// TIA Portal project "Inteligenta_szklarnia" (V15.1) (continued)

screen "tryb_automatyczny" 800x480
   IOField "I/O field_1" at 100,354 size 57x40; FormatPattern 99.9
      ProcessValue <- "Wejscia_HMI_Temperatura"
   Button "Button_1" at 750,0 size 50x50; TextOff 'WRÓĆ'; PictureOff "Back_arrow"
      on Click: function_efd93a16()
   Button "Button_2" at 417,418 size 371x53; TextOff 'ZATWIERDŹ'
      on Click: ActivateScreen("praca", 0)
   Bar "Bar_1" at 14,103 size 70x275; MinimumValue 0; MaximumValue 45
      ProcessValue <- "temperatura_ustawiona_man"
   TextField "Text field_2" at 15,60 size 132x23; Text 'TEMPERATURA'
   Bar "Bar_2" at 217,108 size 70x275; MinimumValue 0; MaximumValue 100
      ProcessValue <- "wilgotnosc_powietrza_man"
   TextField "Text field_3" at 205,61 size 122x42; Text 'WOLGOTNOŚĆ POWIETRZA WILGOTNOŚĆ POWIETRZA'
   Button "Button_3" at 90,119 size 75x45; TextOff '+ / +0.5 °C'
      on Press: function_dd21b452("temperatura_ustawiona_man", 0.5)
   Button "Button_7" at 89,177 size 75x45; TextOff '- / -0.5 °C'
      on Press: function_b9b71300("temperatura_ustawiona_man", 0.5)
   IOField "I/O field_2" at 100,276 size 62x40; FormatPattern 99.9
      ProcessValue <- "temperatura_ustawiona_man"
   TextField "Text field_11" at 155,285 size 23x22; Text '°C'
   TextField "Text field_9" at 155,358 size 23x22; Text '°C'
   Bar "Bar_4" at 417,105 size 70x275; MinimumValue 0; MaximumValue 100
      ProcessValue <- "wilgotnosc_gleby_man"
   TextField "Text field_10" at 404,58 size 122x42; Text 'WOLGOTNOŚĆ GLEBY WILGOTNOŚĆ GLEBY'
   Button "Button_8" at 496,125 size 65x40; TextOff '+ / +2%'
      on Click: function_dd21b452("wilgotnosc_gleby_man", 2)
   Button "Button_9" at 497,177 size 65x40; TextOff '- / -2%'
      on Click: function_b9b71300("wilgotnosc_gleby_man", 2)
   IOField "I/O field_5" at 508,276 size 62x40; FormatPattern 999
      ProcessValue <- "wilgotnosc_gleby_man"
   IOField "I/O field_6" at 508,346 size 62x40; FormatPattern 999
      ProcessValue <- "Parametry_Wilgotność_gleby"
   TextField "Text field_12" at 493,264 size 101x22; Text 'USTAWIONA'
   TextField "Text field_13" at 497,335 size 86x22; Text 'AKTUALNA'
   TextField "Text field_14" at 547,285 size 23x22; Text '%'
   TextField "Text field_15" at 547,356 size 23x22; Text '%'
   Button "Button_10" at 298,125 size 65x40; TextOff '+ / +5%'
      on Click: function_dd21b452("wilgotnosc_powietrza_man", 5)
   Button "Button_11" at 298,177 size 65x40; TextOff '- / -5%'
      on Click: function_b9b71300("wilgotnosc_powietrza_man", 5)
   IOField "I/O field_4" at 305,277 size 66x40; FormatPattern 999
      ProcessValue <- "wilgotnosc_powietrza_man"
   IOField "I/O field_7" at 307,349 size 62x40; FormatPattern 999
      ProcessValue <- "Parametry_Wilgotność_powietrza"
   TextField "Text field_16" at 292,264 size 101x22; Text 'USTAWIONA'
   TextField "Text field_17" at 294,335 size 86x22; Text 'AKTUALNA'
   TextField "Text field_18" at 346,286 size 23x22; Text '%'
   TextField "Text field_19" at 346,357 size 23x22; Text '%'
   Button "Button_14" at 3,1 size 43x43; TextOff 'DOM'; PictureOff "home_1"
      on Click: ActivateScreen("Root screen", 0)
   TextField "Text field_4" at 38,424 size 128x23; Text 'SYSTEM OKIEN'
   Switch "Switch_1" at 198,418 size 185x35; TextOn 'ON'; CaptionText 'Switch'; TextOff 'OFF'
      ProcessValue <- "system_okien"
   GraphicView "Graphic view_1" at 150,60 size 40x40; Picture "Thermometer_icon"
   GraphicView "Graphic view_2" at 330,61 size 40x40; Picture "sensor_4212519"
   TextField "Text field_5" at 93,334 size 86x22; Text 'AKTUALNA'
   TextField "Text field_6" at 90,262 size 101x22; Text 'USTAWIONA'
   GraphicView "Graphic view_3" at 526,61 size 40x40; Picture "soil-sensor_11298794"
   TextField "Text field_1" at 250,4 size 288x34; Text 'TRYB AUTOMATYCZNY'
   Bar "Bar_3" at 620,105 size 70x275; MinimumValue 0; MaximumValue 1500
      ProcessValue <- "wilgotnosc_gleby_man"
   TextField "Text field_7" at 604,53 size 161x42; Text 'WOLGOTNOŚĆ GLEBY NASŁONECZNIENIE'
   GraphicView "Graphic view_4" at 725,79 size 40x40; Picture "sensor_4212513"
   Button "Button_4" at 696,125 size 65x40; TextOff '+ +25 W m'
      on Click: function_dd21b452("naslonecznienie_man", 25)
   Button "Button_5" at 697,177 size 65x40; TextOff '- -25 W m'
      on Click: function_b9b71300("naslonecznienie_man", 25)
   IOField "I/O field_3" at 708,276 size 62x40; FormatPattern 999
      ProcessValue <- "naslonecznienie_man"
   TextField "Text field_8" at 693,264 size 101x22; Text 'USTAWIONA'
   IOField "I/O field_8" at 711,347 size 62x40; FormatPattern 999
      ProcessValue <- "Parametry_Czujnik_światła"
   TextField "Text field_20" at 697,335 size 86x22; Text 'AKTUALNA'
   TextField "Text field_21" at 747,285 size 23x22; Text '%'
   TextField "Text field_22" at 747,356 size 23x22; Text '%'
   TextField "Text field_23" at 751,143 size 32x18; Text '2'
   TextField "Text field_24" at 748,196 size 32x18; Text '2'
*)

(* ===== HMI "HMI_RT_3" =====
system functions are stored by id; their names below are inferred from use
connection "HMI_Connection_4": ETHERNET, SMART_S7_1200_OMS

HMI tags "Default tag table"
   "Tag_ScreenNumber" : UInt, internal

HMI tags "wyjsciaPLC"
   "Alarm_ostrzegwaczy" : Bool = PLC Alarm_ostrzegwaczy AT %Q0.5, 100 ms
   "Grzałka" : Bool = PLC Grzałka AT %Q0.0, 100 ms
   "Pompa_wodna" : Bool = PLC Pompa_wodna AT %Q0.2, 100 ms
   "Rolety_otwieranie" : Bool = PLC Rolety_otwieranie AT %Q0.3, 100 ms
   "Rolety_zamykanie" : Bool = PLC Rolety_zamykanie AT %Q0.4, 100 ms
   "Siłownik_okien_otwieranie" : Bool = PLC Siłownik_okien_otwieranie AT %Q0.6, 100 ms
   "Siłownik_okien_zamykanie" : Bool = PLC Siłownik_okien_zamykanie AT %Q0.7, 100 ms
   "Wentylator" : Bool = PLC Wentylator AT %Q0.1, 100 ms
   "Tag_ScreenNumber(1)" : DInt = PLC Tag_ScreenNumber AT %MD0, 500 ms
   "Parametry_Czujnik_światła" : Int = PLC Parametry.Czujnik_światła, 500 ms
   "Parametry_temeratura" : Real = PLC Parametry.temeratura, 500 ms
   "Parametry_Czujnik_wiatru" : Int = PLC Parametry.Czujnik_wiatru, 500 ms
   "Parametry_Wilgotność_powietrza" : Int = PLC Parametry.Wilgotność_powietrza, 500 ms
   "Parametry_czujnik_CO2" : Int = PLC Parametry.czujnik_CO2, 500 ms
   "Parametry_Wilgotność_gleby" : Int = PLC Parametry.Wilgotność_gleby, 500 ms
   "Wejscia_HMI_Temperatura" : Real = PLC Wejscia_HMI.Temperatura, 500 ms
   "Parametry_stopien_zasloniecia_rolet" : Int = PLC Parametry.stopien_zasloniecia_rolet, 1 s
   "Wejscia_HMI_Zaciemnienie" : Int = PLC Wejscia_HMI.Zaciemnienie, 1 s
   "Receptury_nazwa{0}" : String[254] = PLC Receptury.nazwa[0], 1 s
   "Receptury_nazwa{1}" : String[254] = PLC Receptury.nazwa[1], 1 s
   "Receptury_nazwa{2}" : String[254] = PLC Receptury.nazwa[2], 1 s
   "Receptury_nazwa{3}" : String[254] = PLC Receptury.nazwa[3], 1 s
   "Receptury_nazwa{4}" : String[254] = PLC Receptury.nazwa[4], 1 s
   "Receptury_nazwa{5}" : String[254] = PLC Receptury.nazwa[5], 1 s
   "naslonecznienie_man" : Int = PLC Wejscia_HMI.naslonecznienie_manual, 1 s

HMI tags "USTAWIENIA_HMI"
   "temperatura_ustawiona_man" : Real, internal
   "stopien_otwarcia_okien_man" : Real, internal
   "wilgotnosc_powietrza_man" : Real, internal
   "wilgotnosc_gleby_man" : Real, internal
   "nazwa_receptury" : WString[10], internal
   "system_okien" : Bool, internal
   "AlwaysTRUE" : Bool = PLC AlwaysTRUE AT %M1.2, 1 s

screen "Root screen" 800x480, template "Template_1"
   on GenerateScreen: SetTag("Tag_ScreenNumber", 1)
   Button "Button_3" at 10,270 size 300x90; TextOff 'ZAPISZ NOWĄ RECEPTURĘ'
      on Click: ActivateScreen("zapisz_recepture", 0)
   Button "Button_1" at 10,170 size 300x90; TextOff 'TRYB MANUALNY'
      on Click: ActivateScreen("tryb_manualny", 0)
   Button "Button_2" at 10,70 size 301x90; TextOff 'TRYB AUTOMATYCZNY'
      on Click: ActivateScreen("tryb_automatyczny", 0)
   TextField "Text field_2" at 32,2 size 738x63; Text 'AUTOMATYCZNA SZKLARNIA'
   GraphicView "Graphic view_1" at 370,70 size 392x338; Picture "garden-tools-graphic-clipart-design-free-png"
   Button "Button_4" at 10,370 size 301x90; TextOff 'WYBIERZ RECEPTURĘ'
      on Click: ActivateScreen("wybierz_recepture", 0)
   TextField "Text field_1" at 117,454 size 235x26; Text 'Tego przycisku w symulacji nie widac ale nie chciałem uswac jakby jednak był potrzebny xd'
      Visibility <- "AlwaysTRUE"

screen "zapisz_recepture" 800x480
   TextField "Text field_1" at 282,4 size 253x34; Text 'ZAPISZ RECEPTURE / ZAPISZ RECEPTURĘ'
   Button "Button_1" at 750,0 size 50x50; TextOff 'WRÓĆ'; PictureOff "Back_arrow"
      on Click: function_efd93a16()
   Button "Button_2" at 406,414 size 371x53; TextOff 'ZATWIERDŹ'
      on Click: ActivateScreen("praca", 0)
   Bar "Bar_1" at 17,122 size 70x314; MinimumValue 0; MaximumValue 45
      ProcessValue <- "temperatura_ustawiona_man"
   TextField "Text field_2" at 30,64 size 132x23; Text 'TEMPERATURA'
   Bar "Bar_2" at 223,133 size 54x113; MinimumValue 0; MaximumValue 100
      ProcessValue <- "wilgotnosc_powietrza_man"
   TextField "Text field_3" at 231,45 size 122x42; Text 'WOLGOTNOŚĆ POWIETRZA'
   Button "Button_3" at 115,140 size 73x45; TextOff '+ / +0.5 °C'
      on Press: function_dd21b452("temperatura_ustawiona_man", 0.5)
   Button "Button_7" at 115,201 size 73x45; TextOff '- / -0.5 °C'
      on Press: function_b9b71300("temperatura_ustawiona_man", 0.5)
   TextField "Text field_8" at 93,325 size 109x42; Text 'ustawiona wartość USTAWIONA'
   IOField "I/O field_2" at 106,365 size 62x40; FormatPattern 99.9
      ProcessValue <- "temperatura_ustawiona_man"
   TextField "Text field_11" at 156,367 size 37x37; Text '°C'
   Bar "Bar_4" at 225,346 size 57x127; MinimumValue 0; MaximumValue 100
      ProcessValue <- "wilgotnosc_gleby_man"
   TextField "Text field_10" at 229,254 size 122x42; Text 'WOLGOTNOŚĆ GLEBY'
   Button "Button_8" at 230,300 size 40x40; TextOff '+'
      on Click: function_dd21b452("wilgotnosc_gleby_man", 2)
   Button "Button_9" at 318,300 size 40x40; TextOff '-'
      on Click: function_b9b71300("wilgotnosc_gleby_man", 2)
   IOField "I/O field_5" at 291,401 size 62x40; FormatPattern 999
      ProcessValue <- "wilgotnosc_gleby_man"
   TextField "Text field_12" at 285,384 size 83x20; Text 'USTAWIONA'
   TextField "Text field_14" at 338,404 size 30x29; Text '%'
   Button "Button_10" at 223,87 size 40x40; TextOff '+'
      on Click: function_dd21b452("wilgotnosc_powietrza_man", 5)
   Button "Button_11" at 311,87 size 40x40; TextOff '-'
      on Click: function_b9b71300("wilgotnosc_powietrza_man", 5)
   IOField "I/O field_4" at 291,180 size 62x40; FormatPattern 999
      ProcessValue <- "wilgotnosc_powietrza_man"
   TextField "Text field_16" at 288,167 size 83x20; Text 'USTAWIONA'
   TextField "Text field_18" at 342,184 size 30x29; Text '%'
   Button "Button_14" at 3,1 size 43x43; TextOff 'DOM'; PictureOff "home_1"
      on Click: ActivateScreen("Root screen", 0)
   TextField "Text field_4" at 529,47 size 128x23; Text 'SYSTEM OKIEN'
   Switch "Switch_1" at 503,78 size 185x35; TextOn 'ON'; CaptionText 'Switch'; TextOff 'OFF'
      ProcessValue <- "system_okien"
   IOField "I/O field_1" at 426,311 size 328x81; FormatPattern ????????????????????
      ProcessValue <- "nazwa_receptury"
   TextField "Text field_7" at 406,273 size 380x37; Text 'WPISZ NAZWĘ RECEPTURY'
   GraphicView "Graphic view_1" at 385,338 size 36x30; Picture "Graphic_4"
   GraphicView "Graphic view_2" at 753,338 size 36x30; Picture "Graphic_5"
   TextField "Text field_9" at 387,146 size 161x61; Text 'STOPIEŃ OTWARCIA OKIEN ŚREDNIE NASŁONECZNIENIE'
   Bar "Bar_6" at 404,213 size 373x52; MinimumValue 0; MaximumValue 1500
      ProcessValue <- "naslonecznienie_man"
   Button "Button_4" at 697,145 size 80x50; TextOff '+ / -'
      on Click: function_b9b71300("naslonecznienie_man", 5)
   Button "Button_5" at 589,145 size 80x50; TextOff '- / +'
      on Press: function_dd21b452("naslonecznienie_man", 5)

screen "tryb_manualny" 800x480
   Button "Button_2" at 355,415 size 431x53; TextOff 'ZATWIERDŹ'
      on Click: ActivateScreen("praca", 0)
   TextField "Text field_1" at 282,4 size 223x34; Text 'TRYB MANUALNY'
   Bar "Bar_1" at 181,300 size 60x172; MinimumValue 0; MaximumValue 45
      ProcessValue <- "Parametry_temeratura"
   TextField "Text field_2" at 188,267 size 132x23; Text 'TEMPERATURA'
   Bar "Bar_2" at 181,93 size 60x160; MinimumValue 0; MaximumValue 100
      ProcessValue <- "Parametry_Wilgotność_powietrza"
   TextField "Text field_3" at 198,45 size 122x42; Text 'WOLGOTNOŚĆ POWIETRZA WILGOTNOŚĆ POWIETRZA'
   Bar "Bar_3" at 576,166 size 170x52; MinimumValue 0
      ProcessValue <- "stopien_otwarcia_okien_man"
   TextField "Text field_4" at 576,43 size 186x61; Text 'STOPIEŃ OTWARCIA OKIEN STOPIEŃ OTWARCIA OKIEN'
   IOField "I/O field_1" at 244,368 size 95x40; FormatPattern 99.9
      ProcessValue <- "Wejscia_HMI_Temperatura"
   Bar "Bar_4" at 8,93 size 60x160; MinimumValue 0; MaximumValue 100
      ProcessValue <- "Parametry_Wilgotność_gleby"
   Button "Button_4" at 406,253 size 80x60; TextOff 'PODLEWANIE'
      on Click: InvertBit("Pompa_wodna")
   Button "Button_5" at 536,253 size 80x60; TextOff 'GRZANIE'
      on Click: InvertBit("Grzałka")
   Button "Button_6" at 666,253 size 80x60; TextOff 'WENTYLACJA'
      on Click: InvertBit("Wentylator")
   GraphicView "Graphic view_1" at 675,320 size 60x60; Picture "fan_4829316"
      Visibility <- "Wentylator"
   GraphicView "Graphic view_6" at 545,320 size 60x60; Picture "heater_4463010"
      Visibility <- "Grzałka"
   GraphicView "Graphic view_7" at 415,320 size 60x60; Picture "irrigation_18631825"
      Visibility <- "Pompa_wodna"
   GraphicView "Graphic view_9" at 676,320 size 60x60; Picture "fan_off"
      Visibility <- "Wentylator"
   GraphicView "Graphic view_10" at 546,320 size 60x60; Picture "heater_off"
      Visibility <- "Grzałka"
   GraphicView "Graphic view_11" at 415,320 size 60x60; Picture "irrigation_off"
      Visibility <- "Pompa_wodna"
   TextField "Text field_10" at 18,45 size 122x42; Text 'WOLGOTNOŚĆ GLEBY WILGOTNOŚĆ GLEBY'
   IOField "I/O field_3" at 760,171 size 33x36; FormatPattern 9
      ProcessValue <- "stopien_otwarcia_okien_man"
   IOField "I/O field_6" at 70,148 size 62x40; FormatPattern 999
      ProcessValue <- "Parametry_Wilgotność_gleby"
   TextField "Text field_15" at 115,152 size 35x34; Text '%'
   IOField "I/O field_7" at 252,151 size 62x40; FormatPattern 999
      ProcessValue <- "Parametry_Wilgotność_powietrza"
   TextField "Text field_19" at 294,154 size 35x34; Text '%'
   Button "Button_12" at 576,99 size 50x50; TextOff '+'
      on Click: function_dd21b452("stopien_otwarcia_okien_man", 1)
   Button "Button_13" at 696,98 size 50x50; TextOff '-'
      on Click: function_b9b71300("stopien_otwarcia_okien_man", 1)
   Button "Button_14" at 3,1 size 43x43; TextOff 'DOM'; PictureOff "home_1"
      on Click: ActivateScreen("Root screen", 0)
   Button "Button_1" at 750,0 size 50x50; TextOff 'Text'; PictureOff "Back_arrow"
      on Click: function_efd93a16()
   TextField "Text field_9" at 293,369 size 35x34; Text '°C'
   Circle "Circle_1" at 386,336 size 25x25
      Visibility <- "Pompa_wodna"
   Circle "Circle_4" at 386,336 size 25x25
      Visibility <- "Pompa_wodna"
   Circle "Circle_2" at 511,336 size 25x25
      Visibility <- "Grzałka"
   Circle "Circle_5" at 511,336 size 25x25
      Visibility <- "Grzałka"
   Circle "Circle_3" at 639,336 size 25x25
      Visibility <- "Wentylator"
   Circle "Circle_6" at 639,336 size 25x25
      Visibility <- "Wentylator"
   Bar "Bar_5" at 10,300 size 60x172; MinimumValue 0; MaximumValue 1500
      ProcessValue <- "Parametry_Czujnik_światła"
   TextField "Text field_5" at 3,268 size 161x23; Text 'TEMPERATURA / NASŁONECZNIENIE'
   IOField "I/O field_2" at 70,368 size 95x40; FormatPattern 9999
      ProcessValue <- "Parametry_Czujnik_światła"
   TextField "Text field_6" at 127,356 size 35x64; Text '°C W m'
   TextField "Text field_7" at 152,391 size 31x17; Text '2'
   TextField "Text field_8" at 348,43 size 206x61; Text 'STOPIEŃ OTWARCIA OKIEN STOPIEŃ ZASŁONIENIA ROLET'
   Bar "Bar_6" at 366,166 size 170x52; MinimumValue 0; MaximumValue 100
      ProcessValue <- "naslonecznienie_man"
   Button "Button_3" at 456,98 size 80x50; TextOff '+ / ODSŁOŃ'
      on Click: function_b9b71300("naslonecznienie_man", 5)
   Button "Button_7" at 366,98 size 80x50; TextOff '- / ZASŁOŃ'
      on Press: function_dd21b452("naslonecznienie_man", 5)

screen "wybierz_recepture" 800x480
   TextField "Text field_2" at 257,4 size 280x34; Text 'WYBIERZ RECEPTURE / WYBIERZ RECEPTURĘ'
   Button "Button_1" at 750,0 size 50x50; TextOff 'WRÓĆ'; PictureOff "Back_arrow"
      on Click: function_efd93a16()
   Button "Button_14" at 3,1 size 43x43; TextOff 'DOM'; PictureOff "home_1"
      on Click: ActivateScreen("Root screen", 0)
   TextField "Text field_1" at 18,52 size 23x39; Text '1'
   TextField "Text field_3" at 18,108 size 23x39; Text '2'
   TextField "Text field_4" at 18,169 size 23x39; Text '3'
   TextField "Text field_5" at 18,231 size 23x39; Text '4'
   TextField "Text field_6" at 18,290 size 23x39; Text '5'
   TextField "Text field_7" at 18,351 size 23x39; Text '6'
   Button "Button_2" at 13,415 size 775x55; TextOff '-ZATWIERDŹ-'
      on Click: ActivateScreen("praca", 0)
   Button "Button_3" at 720,68 size 60x60; TextOff 'Text'; PictureOff "Double_up_arrow"
   Button "Button_4" at 720,162 size 60x60; TextOff 'Text'; PictureOff "Double_down_arrow"
   Button "Button_5" at 708,326 size 83x64; TextOff 'USUŃ'
   IOField "I/O field_1" at 90,58 size 243x32; FormatPattern ????????????????????
      ProcessValue <- "Receptury_nazwa{0}"
   IOField "I/O field_2" at 90,115 size 241x32; FormatPattern ????????????????????
      ProcessValue <- "Receptury_nazwa{1}"
   IOField "I/O field_3" at 90,176 size 267x32; FormatPattern ????????????????????
      ProcessValue <- "Receptury_nazwa{2}"
   IOField "I/O field_4" at 90,238 size 264x32; FormatPattern ????????????????????
      ProcessValue <- "Receptury_nazwa{3}"
   IOField "I/O field_5" at 90,294 size 230x32; FormatPattern ????????????????????
      ProcessValue <- "Receptury_nazwa{4}"
   IOField "I/O field_6" at 90,358 size 506x32; FormatPattern ????????????????????
      ProcessValue <- "Receptury_nazwa{5}"

screen "praca" 800x480
   GraphicView "Graphic view_2" at 28,217 size 100x100; Picture "Thermometer_icon"
   GraphicView "Graphic view_4" at 276,362 size 100x100; Picture "soil-sensor_11298794"
   GraphicView "Graphic view_3" at 28,74 size 100x100; Picture "sensor_4212513"
   GraphicView "Graphic view_5" at 276,75 size 100x100; Picture "sensor_4212519"
   GraphicView "Graphic view_1" at 559,362 size 100x100; Picture "fan_4829316"
      Visibility <- "Wentylator"
   GraphicView "Graphic view_6" at 560,217 size 100x100; Picture "heater_4463010"
      Visibility <- "Grzałka"
   GraphicView "Graphic view_7" at 560,75 size 100x100; Picture "irrigation_18631825"
      Visibility <- "Pompa_wodna"
   GraphicView "Graphic view_8" at 28,362 size 100x100; Picture "anemometer_1113716"
   GraphicView "Graphic view_9" at 560,362 size 100x100; Picture "fan_off"
      Visibility <- "Wentylator"
   GraphicView "Graphic view_10" at 561,217 size 100x100; Picture "heater_off"
      Visibility <- "Grzałka"
   GraphicView "Graphic view_11" at 561,75 size 100x100; Picture "irrigation_off"
      Visibility <- "Pompa_wodna"
   GraphicView "Graphic view_12" at 276,217 size 100x100; Picture "sensor_2828470"
   TextField "Text field_1" at 54,52 size 204x23; Text 'INSOLATION / NASŁONECZNIENIE / SONNENEINSTRAHLUNG'
   TextField "Text field_2" at 67,194 size 132x23; Text 'TEMPERATURA'
   TextField "Text field_3" at 46,334 size 166x23; Text 'SZYBKOŚĆ WIATRU'
   TextField "Text field_4" at 349,194 size 123x23; Text 'STĘŻENIE CO2'
   TextField "Text field_5" at 294,50 size 223x23; Text 'WILGOTNOŚĆ POWIETRZA'
   TextField "Text field_6" at 321,339 size 175x23; Text 'WILGOTNOŚĆ GLEBY'
   TextField "Text field_7" at 626,46 size 116x23; Text 'PODLEWANIE'
   TextField "Text field_8" at 643,192 size 80x23; Text 'GRZANIE'
   TextField "Text field_9" at 626,330 size 117x23; Text 'WENTYLACJA'
   TextField "Text field_10" at 282,4 size 256x34; Text 'PODGLĄD NA ŻYWO'
   Button "Button_1" at 750,0 size 50x50; TextOff 'WRÓĆ'; PictureOff "Back_arrow"
      on Click: function_efd93a16()
   Button "Button_2" at 3,1 size 43x43; TextOff 'DOM'; PictureOff "home_1"
      on Click: ActivateScreen("Root screen", 0)
   IOField "I/O field_2" at 120,233 size 97x65; FormatPattern 99.99
      ProcessValue <- "Parametry_temeratura"
   IOField "I/O field_3" at 136,383 size 70x65; FormatPattern 999
      ProcessValue <- "Parametry_Czujnik_wiatru"
   IOField "I/O field_5" at 377,235 size 83x65; FormatPattern 9999
      ProcessValue <- "Parametry_czujnik_CO2"
   TextField "Text field_11" at 214,241 size 46x46; Text '°C'
   IOField "I/O field_4" at 406,95 size 69x65; FormatPattern 999
      ProcessValue <- "Parametry_Wilgotność_powietrza"
   IOField "I/O field_6" at 406,384 size 68x65; FormatPattern 999
      ProcessValue <- "Parametry_Wilgotność_gleby"
   TextField "Text field_12" at 472,106 size 47x46; Text '%'
   TextField "Text field_13" at 472,396 size 47x46; Text '%'
   TextField "Text field_14" at 219,90 size 47x72; Text 'W m²'
   IOField "I/O field_1" at 119,109 size 101x32; FormatPattern 99999
      ProcessValue <- "Parametry_Czujnik_światła"
   TextField "Text field_15" at 210,376 size 52x72; Text 'Km h'
   Circle "Circle_1" at 695,101 size 48x48
      Visibility <- "Pompa_wodna"
   Circle "Circle_2" at 695,243 size 48x48
      Visibility <- "Grzałka"
   TextField "Text field_16" at 472,242 size 69x39; Text 'ppm'
   Circle "Circle_4" at 695,101 size 48x48
      Visibility <- "Pompa_wodna"
   Circle "Circle_5" at 695,243 size 48x48
      Visibility <- "Grzałka"
   Circle "Circle_3" at 695,385 size 48x48
      Visibility <- "Wentylator"
   Circle "Circle_6" at 695,385 size 48x48
      Visibility <- "Wentylator"

screen "tryb_automatyczny" 800x480
   IOField "I/O field_1" at 100,354 size 57x40; FormatPattern 99.9
      ProcessValue <- "Wejscia_HMI_Temperatura"
   Button "Button_1" at 750,0 size 50x50; TextOff 'WRÓĆ'; PictureOff "Back_arrow"
      on Click: function_efd93a16()
   Button "Button_2" at 417,418 size 371x53; TextOff 'ZATWIERDŹ'
      on Click: ActivateScreen("praca", 0)
   Bar "Bar_1" at 14,103 size 70x275; MinimumValue 0; MaximumValue 45
      ProcessValue <- "temperatura_ustawiona_man"
   TextField "Text field_2" at 15,60 size 132x23; Text 'TEMPERATURA'
   Bar "Bar_2" at 217,108 size 70x275; MinimumValue 0; MaximumValue 100
      ProcessValue <- "wilgotnosc_powietrza_man"
   TextField "Text field_3" at 205,61 size 122x42; Text 'WOLGOTNOŚĆ POWIETRZA WILGOTNOŚĆ POWIETRZA'
   Button "Button_3" at 90,119 size 75x45; TextOff '+ / +0.5 °C'
      on Press: function_dd21b452("temperatura_ustawiona_man", 0.5)
   Button "Button_7" at 89,177 size 75x45; TextOff '- / -0.5 °C'
      on Press: function_b9b71300("temperatura_ustawiona_man", 0.5)
   IOField "I/O field_2" at 100,276 size 62x40; FormatPattern 99.9
      ProcessValue <- "temperatura_ustawiona_man"
   TextField "Text field_11" at 155,285 size 23x22; Text '°C'
   TextField "Text field_9" at 155,358 size 23x22; Text '°C'
   Bar "Bar_4" at 417,105 size 70x275; MinimumValue 0; MaximumValue 100
      ProcessValue <- "wilgotnosc_gleby_man"
   TextField "Text field_10" at 404,58 size 122x42; Text 'WOLGOTNOŚĆ GLEBY WILGOTNOŚĆ GLEBY'
   Button "Button_8" at 496,125 size 65x40; TextOff '+ / +2%'
      on Click: function_dd21b452("wilgotnosc_gleby_man", 2)
   Button "Button_9" at 497,177 size 65x40; TextOff '- / -2%'
      on Click: function_b9b71300("wilgotnosc_gleby_man", 2)
   IOField "I/O field_5" at 508,276 size 62x40; FormatPattern 999
      ProcessValue <- "wilgotnosc_gleby_man"
   IOField "I/O field_6" at 508,346 size 62x40; FormatPattern 999
      ProcessValue <- "Parametry_Wilgotność_gleby"
   TextField "Text field_12" at 493,264 size 101x22; Text 'USTAWIONA'
   TextField "Text field_13" at 497,335 size 86x22; Text 'AKTUALNA'
   TextField "Text field_14" at 547,285 size 23x22; Text '%'
   TextField "Text field_15" at 547,356 size 23x22; Text '%'
   Button "Button_10" at 298,125 size 65x40; TextOff '+ / +5%'
      on Click: function_dd21b452("wilgotnosc_powietrza_man", 5)
   Button "Button_11" at 298,177 size 65x40; TextOff '- / -5%'
      on Click: function_b9b71300("wilgotnosc_powietrza_man", 5)
   IOField "I/O field_4" at 305,277 size 66x40; FormatPattern 999
      ProcessValue <- "wilgotnosc_powietrza_man"
   IOField "I/O field_7" at 307,349 size 62x40; FormatPattern 999
      ProcessValue <- "Parametry_Wilgotność_powietrza"
   TextField "Text field_16" at 292,264 size 101x22; Text 'USTAWIONA'
   TextField "Text field_17" at 294,335 size 86x22; Text 'AKTUALNA'
   TextField "Text field_18" at 346,286 size 23x22; Text '%'
   TextField "Text field_19" at 346,357 size 23x22; Text '%'
   Button "Button_14" at 3,1 size 43x43; TextOff 'DOM'; PictureOff "home_1"
      on Click: ActivateScreen("Root screen", 0)
   TextField "Text field_4" at 38,424 size 128x23; Text 'SYSTEM OKIEN'
   Switch "Switch_1" at 198,418 size 185x35; TextOn 'ON'; CaptionText 'Switch'; TextOff 'OFF'
      ProcessValue <- "system_okien"
   GraphicView "Graphic view_1" at 150,60 size 40x40; Picture "Thermometer_icon"
   GraphicView "Graphic view_2" at 330,61 size 40x40; Picture "sensor_4212519"
   TextField "Text field_5" at 93,334 size 86x22; Text 'AKTUALNA'
   TextField "Text field_6" at 90,262 size 101x22; Text 'USTAWIONA'
   GraphicView "Graphic view_3" at 526,61 size 40x40; Picture "soil-sensor_11298794"
   TextField "Text field_1" at 250,4 size 288x34; Text 'TRYB AUTOMATYCZNY'
   Bar "Bar_3" at 620,105 size 70x275; MinimumValue 0; MaximumValue 1500
      ProcessValue <- "wilgotnosc_gleby_man"
   TextField "Text field_7" at 604,53 size 161x42; Text 'WOLGOTNOŚĆ GLEBY NASŁONECZNIENIE'
   GraphicView "Graphic view_4" at 725,79 size 40x40; Picture "sensor_4212513"
   Button "Button_4" at 696,125 size 65x40; TextOff '+ +25 W m'
      on Click: function_dd21b452("naslonecznienie_man", 25)
   Button "Button_5" at 697,177 size 65x40; TextOff '- -25 W m'
      on Click: function_b9b71300("naslonecznienie_man", 25)
   IOField "I/O field_3" at 708,276 size 62x40; FormatPattern 999
      ProcessValue <- "naslonecznienie_man"
   TextField "Text field_8" at 693,264 size 101x22; Text 'USTAWIONA'
   IOField "I/O field_8" at 711,347 size 62x40; FormatPattern 999
      ProcessValue <- "Parametry_Czujnik_światła"
   TextField "Text field_20" at 697,335 size 86x22; Text 'AKTUALNA'
   TextField "Text field_21" at 747,285 size 23x22; Text '%'
   TextField "Text field_22" at 747,356 size 23x22; Text '%'
   TextField "Text field_23" at 751,143 size 32x18; Text '2'
   TextField "Text field_24" at 748,196 size 32x18; Text '2'

Template "Template_1" 800x480
   Button "Exit" at 671,429 size 71x50; TextOn 'Exit'; TextOff 'Exit'; PictureOn "ExitRuntime_KTP700_Basic_PN_TR"; PictureOff "ExitRuntime_KTP700_Basic_PN_TR"
      on Release: StopRuntime(0)
   Button "Alarms" at 524,429 size 71x50; TextOn 'Alarms'; TextOff 'Alarms'; PictureOn "AlarmDisplay_KTP700_Basic_PN_TR"; PictureOff "AlarmDisplay_KTP700_Basic_PN_TR"
      on Release: function_ef3f5d25("Alarm window_Unacknowledged", -1)
   Button "Start screen" at 169,429 size 71x50; TextOn 'Start screen'; TextOff 'Start screen'; PictureOn "NavigateHome_KTP700_Basic_PN_TR"; PictureOff "NavigateHome_KTP700_Basic_PN_TR"
      on Release: ActivateScreen("Root screen", 0)
      Visibility <- "AlwaysTRUE"
   Button "Language" at 377,429 size 71x50; TextOn 'Language'; TextOff 'Language'; PictureOn "ToggleLanguage_KTP700_Basic_PN_TR"; PictureOff "ToggleLanguage_KTP700_Basic_PN_TR"
      on Release: function_fb9197e8(-1)
*)

(* ===== HMI "HMI_RT_2" =====
system functions are stored by id; their names below are inferred from use
connection "HMI_Connection_3": ETHERNET, SMART_S7_1200_OMS

HMI tags "Default tag table"
   "Tag_ScreenNumber" : Int = PLC HMI.Numer_ekranu_HMI AT %MD0, 500 ms
   "AlwaysTRUE" : Bool = PLC AlwaysTRUE AT %M1.2, 1 s

HMI tags "Receptury"
   "Receptury_nazwa{0}" : String[254] = PLC Receptury.nazwa[0], 1 s
   "Receptury_nazwa{1}" : String[254] = PLC Receptury.nazwa[1], 1 s
   "Receptury_nazwa{2}" : String[254] = PLC Receptury.nazwa[2], 1 s
   "Receptury_nazwa{3}" : String[254] = PLC Receptury.nazwa[3], 1 s
   "Receptury_nazwa{4}" : String[254] = PLC Receptury.nazwa[4], 1 s
   "Receptury_nazwa{5}" : String[254] = PLC Receptury.nazwa[5], 1 s

HMI tags "USTAWIENIA_HMI"
   "nazwa_receptury" : WString[10], internal

HMI tags "Do_PLC"
   "System_okien_auto" : Bool = PLC HMI.System_okien_auto, 500 ms
   "Stopien_zasloniecia_rolet_manual" : Int = PLC HMI.Stopien_zasloniecia_rolet_manual, 100 ms
   "Przycisk_pompy_manual" : Bool = PLC HMI.Przycisk_pompa_manual AT %Q0.2, 100 ms
   "Przycisk_wentylacja_manual" : Bool = PLC HMI.Przycisk_wentylacja_manual AT %Q0.1, 100 ms
   "Przycisk_grzanie_manual" : Bool = PLC HMI.Przycisk_grzanie_manual AT %Q0.0, 100 ms
   "Stopien_otwarcia_okien_man" : Int = PLC HMI.Stopien_otwarcia_okien_manual AT %DB1.DBW0, 100 ms
   "Temperatura_auto" : Real = PLC HMI.Temperatura_auto, 500 ms
   "Naslonecznienie_auto" : Int = PLC HMI.Naslonecznienie_auto AT %DB1.DBW0, 500 ms
   "Wilgotnosc_powietrza_auto" : Int = PLC HMI.Wilgotnosc_powietrza_auto AT %DB1.DBW0, 500 ms
   "Wilgotnosc_gleby_auto" : Int = PLC HMI.Wilgotnosc_gleby_auto AT %DB1.DBW0, 500 ms
   "Przycisk_zatwierdz" : Bool = PLC HMI.Przycisk_zatwierdz AT %DB1.DBW0, 100 ms

HMI tags "Z_PLC"
   "Czujnik_wilgotności_powietrza" : Int = PLC Wejscia_PLC.Czujnik_wilgotności_powietrza, 500 ms
   "Czujnik_temeratury_wewnetrznej" : Real = PLC Wejscia_PLC.Temeratura_wewnetrzna, 500 ms
   "Czujnik_natezenia_światła" : Int = PLC Wejscia_PLC.Czujnik_natezenia_swiatła, 500 ms
   "Czujnik_wilgotności_gleby" : Int = PLC Wejscia_PLC.Czujnik_wilgotności_gleby, 500 ms
   "Czujnik_CO2" : Int = PLC Wejscia_PLC.Czujnik_CO2, 500 ms
   "Czujnik_wiatru" : Int = PLC Wejscia_PLC.Czujnik_wiatru, 500 ms
   "Stopien_zasloniecia_rolet" : Int = PLC Wejscia_PLC.Stopien_zasloniecia_rolet, 1 s

screen "Root screen" 800x480, template "Template_1"
   on GenerateScreen: SetTag("Tag_ScreenNumber", 0)
   Button "Button_3" at 10,270 size 300x90; TextOff 'ZAPISZ NOWĄ RECEPTURĘ'
      on Click: ActivateScreen("zapisz_recepture", 0)
   Button "Button_1" at 10,170 size 300x90; TextOff 'TRYB MANUALNY'
      on Click: ActivateScreen("tryb_manualny", 0)
   Button "Button_2" at 10,70 size 301x90; TextOff 'TRYB AUTOMATYCZNY'
      on Click: ActivateScreen("tryb_automatyczny", 0)
   TextField "Text field_2" at 32,2 size 738x63; Text 'AUTOMATYCZNA SZKLARNIA'
   GraphicView "Graphic view_1" at 370,70 size 392x338; Picture "garden-tools-graphic-clipart-design-free-png"
   Button "Button_4" at 10,370 size 301x90; TextOff 'WYBIERZ RECEPTURĘ'
      on Click: ActivateScreen("wybierz_recepture", 0)

screen "zapisz_recepture" 800x480
   on GenerateScreen: SetTag("Tag_ScreenNumber", 4)
   TextField "Text field_1" at 282,4 size 253x34; Text 'ZAPISZ RECEPTURE / ZAPISZ RECEPTURĘ'
   Button "Button_1" at 750,0 size 50x50; TextOff 'WRÓĆ'; PictureOff "Back_arrow"
      on Click: function_efd93a16()
   Button "Button_2" at 406,414 size 371x53; TextOff 'ZATWIERDŹ'
      on Click: ActivateScreen("praca", 0)
      on Press: function_b14e0dd5("Przycisk_zatwierdz", 0)
   Bar "Bar_1" at 17,122 size 70x314; MinimumValue 0; MaximumValue 45
      ProcessValue <- "Temperatura_auto"
   TextField "Text field_2" at 30,64 size 132x23; Text 'TEMPERATURA'
   Bar "Bar_2" at 223,133 size 54x113; MinimumValue 0; MaximumValue 100
      ProcessValue <- "Wilgotnosc_powietrza_auto"
   TextField "Text field_3" at 231,45 size 122x42; Text 'WOLGOTNOŚĆ POWIETRZA'
   Button "Button_3" at 115,140 size 73x45; TextOff '+ / +0.5 °C'
      on Press: function_dd21b452("Temperatura_auto", 0.5)
   Button "Button_7" at 115,201 size 73x45; TextOff '- / -0.5 °C'
      on Press: function_b9b71300("Temperatura_auto", 0.5)
   TextField "Text field_8" at 93,325 size 109x42; Text 'ustawiona wartość USTAWIONA'
   IOField "I/O field_2" at 106,365 size 62x40; FormatPattern 99.9
      ProcessValue <- "Temperatura_auto"
   TextField "Text field_11" at 156,367 size 37x37; Text '°C'
   Bar "Bar_4" at 225,346 size 57x127; MinimumValue 0; MaximumValue 100
      ProcessValue <- "Wilgotnosc_gleby_auto"
   TextField "Text field_10" at 229,254 size 122x42; Text 'WOLGOTNOŚĆ GLEBY'
   Button "Button_8" at 230,300 size 40x40; TextOff '+'
      on Click: function_dd21b452("Wilgotnosc_gleby_auto", 2)
   Button "Button_9" at 318,300 size 40x40; TextOff '-'
      on Click: function_b9b71300("Wilgotnosc_gleby_auto", 2)
   IOField "I/O field_5" at 291,401 size 62x40; FormatPattern 999
      ProcessValue <- "Wilgotnosc_gleby_auto"
   TextField "Text field_12" at 285,384 size 83x20; Text 'USTAWIONA'
   TextField "Text field_14" at 338,404 size 30x29; Text '%'
   Button "Button_10" at 223,87 size 40x40; TextOff '+'
      on Click: function_dd21b452("Wilgotnosc_powietrza_auto", 5)
   Button "Button_11" at 311,87 size 40x40; TextOff '-'
      on Click: function_b9b71300("Wilgotnosc_powietrza_auto", 5)
   IOField "I/O field_4" at 291,180 size 62x40; FormatPattern 999
      ProcessValue <- "Wilgotnosc_powietrza_auto"
   TextField "Text field_16" at 288,167 size 83x20; Text 'USTAWIONA'
   TextField "Text field_18" at 342,184 size 30x29; Text '%'
   Button "Button_14" at 3,1 size 43x43; TextOff 'DOM'; PictureOff "home_1"
      on Click: ActivateScreen("Root screen", 0)
   TextField "Text field_4" at 529,47 size 128x23; Text 'SYSTEM OKIEN'
   Switch "Switch_1" at 503,78 size 185x35; TextOn 'ON'; CaptionText 'Switch'; TextOff 'OFF'
      ProcessValue <- "System_okien_auto"
   IOField "I/O field_1" at 426,311 size 328x81; FormatPattern ????????????????????
      ProcessValue <- "nazwa_receptury"
   TextField "Text field_7" at 406,273 size 380x37; Text 'WPISZ NAZWĘ RECEPTURY'
   GraphicView "Graphic view_1" at 385,338 size 36x30; Picture "Graphic_4"
   GraphicView "Graphic view_2" at 753,338 size 36x30; Picture "Graphic_5"
   TextField "Text field_9" at 387,146 size 161x61; Text 'STOPIEŃ OTWARCIA OKIEN ŚREDNIE NASŁONECZNIENIE'
   Bar "Bar_6" at 404,213 size 373x52; MinimumValue 0; MaximumValue 1500
      ProcessValue <- "Stopien_zasloniecia_rolet_manual"
   Button "Button_4" at 697,145 size 80x50; TextOff '+ / -'
      on Click: function_b9b71300("Stopien_zasloniecia_rolet_manual", 5)
   Button "Button_5" at 589,145 size 80x50; TextOff '- / +'
      on Press: function_dd21b452("Stopien_zasloniecia_rolet_manual", 5)

screen "tryb_manualny" 800x480
   on GenerateScreen: SetTag("Tag_ScreenNumber", 2)
   TextField "Text field_1" at 282,4 size 223x34; Text 'TRYB MANUALNY'
   Bar "Bar_1" at 181,300 size 60x172; MinimumValue 0; MaximumValue 45
      ProcessValue <- "Czujnik_temeratury_wewnetrznej"
   TextField "Text field_2" at 188,267 size 132x23; Text 'TEMPERATURA'
   Bar "Bar_2" at 181,93 size 60x160; MinimumValue 0; MaximumValue 100
      ProcessValue <- "Czujnik_wilgotności_powietrza"
   TextField "Text field_3" at 198,45 size 122x42; Text 'WOLGOTNOŚĆ POWIETRZA WILGOTNOŚĆ POWIETRZA'
   Bar "Bar_3" at 576,166 size 170x52; MinimumValue 0
      ProcessValue <- "Stopien_otwarcia_okien_man"
   TextField "Text field_4" at 576,43 size 186x61; Text 'STOPIEŃ OTWARCIA OKIEN STOPIEŃ OTWARCIA OKIEN'
   IOField "I/O field_1" at 244,368 size 95x40; FormatPattern 99.9
      ProcessValue <- "Czujnik_temeratury_wewnetrznej"
   Bar "Bar_4" at 8,93 size 60x160; MinimumValue 0; MaximumValue 100
      ProcessValue <- "Czujnik_wilgotności_gleby"
   Button "Button_4" at 380,253 size 97x80; TextOff 'PODLEWANIE'
      on Click: InvertBit("Przycisk_pompy_manual")
   Button "Button_5" at 522,253 size 100x80; TextOff 'GRZANIE'
      on Click: InvertBit("Przycisk_grzanie_manual")
   Button "Button_6" at 671,253 size 100x80; TextOff 'WENTYLACJA'
      on Click: InvertBit("Przycisk_wentylacja_manual")
   GraphicView "Graphic view_1" at 681,356 size 76x80; Picture "fan_4829316"
      Visibility <- "Przycisk_wentylacja_manual"
   GraphicView "Graphic view_6" at 529,356 size 80x80; Picture "heater_4463010"
      Visibility <- "Przycisk_grzanie_manual"
   GraphicView "Graphic view_7" at 394,356 size 77x80; Picture "irrigation_18631825"
      Visibility <- "Przycisk_pompy_manual"
   GraphicView "Graphic view_9" at 682,356 size 76x80; Picture "fan_off"
      Visibility <- "Przycisk_wentylacja_manual"
   GraphicView "Graphic view_10" at 530,356 size 80x80; Picture "heater_off"
      Visibility <- "Przycisk_grzanie_manual"
   GraphicView "Graphic view_11" at 394,356 size 77x80; Picture "irrigation_off"
      Visibility <- "Przycisk_pompy_manual"
   TextField "Text field_10" at 18,45 size 122x42; Text 'WOLGOTNOŚĆ GLEBY WILGOTNOŚĆ GLEBY'
   IOField "I/O field_3" at 760,171 size 33x36; FormatPattern 9
      ProcessValue <- "Stopien_otwarcia_okien_man"
   IOField "I/O field_6" at 70,148 size 62x40; FormatPattern 999
      ProcessValue <- "Czujnik_wilgotności_gleby"
   TextField "Text field_15" at 115,152 size 35x34; Text '%'
   IOField "I/O field_7" at 252,151 size 62x40; FormatPattern 999
      ProcessValue <- "Czujnik_wilgotności_powietrza"
   TextField "Text field_19" at 294,154 size 35x34; Text '%'
   Button "Button_12" at 576,99 size 50x50; TextOff '+'
      on Click: function_dd21b452("Stopien_otwarcia_okien_man", 1)
   Button "Button_13" at 696,98 size 50x50; TextOff '-'
      on Click: function_b9b71300("Stopien_otwarcia_okien_man", 1)
   Button "Button_14" at 3,1 size 43x43; TextOff 'DOM'; PictureOff "home_1"
      on Click: ActivateScreen("Root screen", 0)
   Button "Button_1" at 750,0 size 50x50; TextOff 'Text'; PictureOff "Back_arrow"
      on Click: function_efd93a16()
   TextField "Text field_9" at 293,369 size 35x34; Text '°C'
   Circle "Circle_1" at 352,378 size 42x42
      Visibility <- "Przycisk_pompy_manual"
   Circle "Circle_4" at 352,378 size 42x42
      Visibility <- "Przycisk_pompy_manual"
   Circle "Circle_2" at 486,375 size 42x42
      Visibility <- "Przycisk_grzanie_manual"
   Circle "Circle_5" at 486,375 size 42x42
      Visibility <- "Przycisk_grzanie_manual"
   Circle "Circle_3" at 630,375 size 41x41
      Visibility <- "Przycisk_wentylacja_manual"
   Circle "Circle_6" at 630,375 size 41x41
      Visibility <- "Przycisk_wentylacja_manual"
   Bar "Bar_5" at 10,300 size 60x172; MinimumValue 0; MaximumValue 1500
      ProcessValue <- "Czujnik_natezenia_światła"
   TextField "Text field_5" at 3,268 size 161x23; Text 'TEMPERATURA / NASŁONECZNIENIE'
   IOField "I/O field_2" at 70,368 size 95x40; FormatPattern 9999
      ProcessValue <- "Czujnik_natezenia_światła"
   TextField "Text field_6" at 127,356 size 35x64; Text '°C W m'
   TextField "Text field_7" at 152,391 size 31x17; Text '2'
   TextField "Text field_8" at 348,43 size 205x61; Text 'STOPIEŃ OTWARCIA OKIEN STOPIEŃ ZASŁONIECIA ROLET'
   Bar "Bar_6" at 366,166 size 170x52; MinimumValue 0; MaximumValue 100
      ProcessValue <- "Stopien_zasloniecia_rolet_manual"
   Button "Button_3" at 456,98 size 80x50; TextOff '+ / ODSŁOŃ'
      on Click: function_b9b71300("Stopien_zasloniecia_rolet_manual", 5)
   Button "Button_7" at 366,98 size 80x50; TextOff '- / ZASŁOŃ'
      on Press: function_dd21b452("Stopien_zasloniecia_rolet_manual", 5)

screen "wybierz_recepture" 800x480
   on GenerateScreen: SetTag("Tag_ScreenNumber", 3)
   TextField "Text field_2" at 257,4 size 280x34; Text 'WYBIERZ RECEPTURE / WYBIERZ RECEPTURĘ'
   Button "Button_1" at 750,0 size 50x50; TextOff 'WRÓĆ'; PictureOff "Back_arrow"
      on Click: function_efd93a16()
   Button "Button_14" at 3,1 size 43x43; TextOff 'DOM'; PictureOff "home_1"
      on Click: ActivateScreen("Root screen", 0)
   TextField "Text field_1" at 18,52 size 23x39; Text '1'
   TextField "Text field_3" at 18,108 size 23x39; Text '2'
   TextField "Text field_4" at 18,169 size 23x39; Text '3'
   TextField "Text field_5" at 18,231 size 23x39; Text '4'
   TextField "Text field_6" at 18,290 size 23x39; Text '5'
   TextField "Text field_7" at 18,351 size 23x39; Text '6'
   Button "Button_2" at 13,415 size 775x55; TextOff '-ZATWIERDŹ-'
      on Click: ActivateScreen("praca", 0)
      on Press: function_b14e0dd5("Przycisk_zatwierdz", 0)
   Button "Button_3" at 720,68 size 60x60; TextOff 'Text'; PictureOff "Double_up_arrow"
   Button "Button_4" at 720,162 size 60x60; TextOff 'Text'; PictureOff "Double_down_arrow"
   Button "Button_5" at 708,326 size 83x64; TextOff 'USUŃ'
   IOField "I/O field_1" at 90,58 size 243x32; FormatPattern ????????????????????
      ProcessValue <- "Receptury_nazwa{0}"
   IOField "I/O field_2" at 90,115 size 241x32; FormatPattern ????????????????????
      ProcessValue <- "Receptury_nazwa{1}"
   IOField "I/O field_3" at 90,176 size 267x32; FormatPattern ????????????????????
      ProcessValue <- "Receptury_nazwa{2}"
   IOField "I/O field_4" at 90,238 size 264x32; FormatPattern ????????????????????
      ProcessValue <- "Receptury_nazwa{3}"
   IOField "I/O field_5" at 90,294 size 230x32; FormatPattern ????????????????????
      ProcessValue <- "Receptury_nazwa{4}"
   IOField "I/O field_6" at 90,358 size 506x32; FormatPattern ????????????????????
      ProcessValue <- "Receptury_nazwa{5}"

screen "praca" 800x480
   on GenerateScreen: SetTag("Tag_ScreenNumber", 5)
   GraphicView "Graphic view_2" at 28,217 size 100x100; Picture "Thermometer_icon"
   GraphicView "Graphic view_4" at 276,362 size 100x100; Picture "soil-sensor_11298794"
   GraphicView "Graphic view_3" at 28,74 size 100x100; Picture "sensor_4212513"
   GraphicView "Graphic view_5" at 276,75 size 100x100; Picture "sensor_4212519"
   GraphicView "Graphic view_1" at 559,362 size 100x100; Picture "fan_4829316"
      Visibility <- "Przycisk_wentylacja_manual"
   GraphicView "Graphic view_6" at 560,217 size 100x100; Picture "heater_4463010"
      Visibility <- "Przycisk_grzanie_manual"
   GraphicView "Graphic view_7" at 560,75 size 100x100; Picture "irrigation_18631825"
      Visibility <- "Przycisk_pompy_manual"
   GraphicView "Graphic view_8" at 28,362 size 100x100; Picture "anemometer_1113716"
   GraphicView "Graphic view_9" at 560,362 size 100x100; Picture "fan_off"
      Visibility <- "Przycisk_wentylacja_manual"
   GraphicView "Graphic view_10" at 561,217 size 100x100; Picture "heater_off"
      Visibility <- "Przycisk_grzanie_manual"
   GraphicView "Graphic view_11" at 561,75 size 100x100; Picture "irrigation_off"
      Visibility <- "Przycisk_pompy_manual"
   GraphicView "Graphic view_12" at 276,217 size 100x100; Picture "sensor_2828470"
   TextField "Text field_1" at 54,52 size 204x23; Text 'INSOLATION / NASŁONECZNIENIE / SONNENEINSTRAHLUNG'
   TextField "Text field_2" at 67,194 size 132x23; Text 'TEMPERATURA'
   TextField "Text field_3" at 46,334 size 166x23; Text 'SZYBKOŚĆ WIATRU'
   TextField "Text field_4" at 349,194 size 123x23; Text 'STĘŻENIE CO2'
   TextField "Text field_5" at 294,50 size 223x23; Text 'WILGOTNOŚĆ POWIETRZA'
   TextField "Text field_6" at 321,339 size 175x23; Text 'WILGOTNOŚĆ GLEBY'
   TextField "Text field_7" at 626,46 size 116x23; Text 'PODLEWANIE'
   TextField "Text field_8" at 643,192 size 80x23; Text 'GRZANIE'
   TextField "Text field_9" at 626,330 size 117x23; Text 'WENTYLACJA'
   TextField "Text field_10" at 282,4 size 256x34; Text 'PODGLĄD NA ŻYWO'
   Button "Button_1" at 750,0 size 50x50; TextOff 'WRÓĆ'; PictureOff "Back_arrow"
      on Click: function_efd93a16()
   Button "Button_2" at 3,1 size 43x43; TextOff 'DOM'; PictureOff "home_1"
      on Click: ActivateScreen("Root screen", 0)
   IOField "I/O field_2" at 120,233 size 97x65; FormatPattern 99.99
      ProcessValue <- "Czujnik_temeratury_wewnetrznej"
   IOField "I/O field_3" at 136,383 size 70x65; FormatPattern 999
      ProcessValue <- "Czujnik_wiatru"
   IOField "I/O field_5" at 377,235 size 83x65; FormatPattern 9999
      ProcessValue <- "Czujnik_CO2"
   TextField "Text field_11" at 214,241 size 46x46; Text '°C'
   IOField "I/O field_4" at 406,95 size 69x65; FormatPattern 999
      ProcessValue <- "Czujnik_wilgotności_powietrza"
   IOField "I/O field_6" at 406,384 size 68x65; FormatPattern 999
      ProcessValue <- "Czujnik_wilgotności_gleby"
   TextField "Text field_12" at 472,106 size 47x46; Text '%'
   TextField "Text field_13" at 472,396 size 47x46; Text '%'
   TextField "Text field_14" at 219,90 size 47x72; Text 'W m²'
   IOField "I/O field_1" at 119,109 size 101x32; FormatPattern 99999
      ProcessValue <- "Czujnik_natezenia_światła"
   TextField "Text field_15" at 210,376 size 52x72; Text 'Km h'
   Circle "Circle_1" at 695,101 size 48x48
      Visibility <- "Przycisk_pompy_manual"
   Circle "Circle_2" at 695,243 size 48x48
      Visibility <- "Przycisk_grzanie_manual"
   TextField "Text field_16" at 472,242 size 69x39; Text 'ppm'
   Circle "Circle_4" at 695,101 size 48x48
      Visibility <- "Przycisk_pompy_manual"
   Circle "Circle_5" at 695,243 size 48x48
      Visibility <- "Przycisk_grzanie_manual"
   Circle "Circle_3" at 695,385 size 48x48
      Visibility <- "Przycisk_wentylacja_manual"
   Circle "Circle_6" at 695,385 size 48x48
      Visibility <- "Przycisk_wentylacja_manual"

screen "tryb_automatyczny" 800x480
   on GenerateScreen: SetTag("Tag_ScreenNumber", 1)
   IOField "I/O field_1" at 100,354 size 57x40; FormatPattern 99.9
      ProcessValue <- "Czujnik_temeratury_wewnetrznej"
   Button "Button_1" at 750,0 size 50x50; TextOff 'WRÓĆ'; PictureOff "Back_arrow"
      on Click: function_efd93a16()
   Button "Button_2" at 417,418 size 371x53; TextOff 'ZATWIERDŹ'
      on Click: ActivateScreen("praca", 0)
      on Press: function_b14e0dd5("Przycisk_zatwierdz", 0)
   Bar "Bar_1" at 14,103 size 70x275; MinimumValue 0; MaximumValue 45
      ProcessValue <- "Temperatura_auto"
   TextField "Text field_2" at 15,60 size 132x23; Text 'TEMPERATURA'
   Bar "Bar_2" at 217,108 size 70x275; MinimumValue 0; MaximumValue 100
      ProcessValue <- "Wilgotnosc_powietrza_auto"
   TextField "Text field_3" at 205,61 size 122x42; Text 'WOLGOTNOŚĆ POWIETRZA WILGOTNOŚĆ POWIETRZA'
   Button "Button_3" at 90,119 size 75x45; TextOff '+ / +0.5 °C'
      on Press: function_dd21b452("Temperatura_auto", 0.5)
   Button "Button_7" at 89,177 size 75x45; TextOff '- / -0.5 °C'
      on Press: function_b9b71300("Temperatura_auto", 0.5)
   IOField "I/O field_2" at 100,276 size 62x40; FormatPattern 99.9
      ProcessValue <- "Temperatura_auto"
   TextField "Text field_11" at 155,285 size 23x22; Text '°C'
   TextField "Text field_9" at 155,358 size 23x22; Text '°C'
   Bar "Bar_4" at 417,105 size 70x275; MinimumValue 0; MaximumValue 100
      ProcessValue <- "Wilgotnosc_gleby_auto"
   TextField "Text field_10" at 404,58 size 122x42; Text 'WOLGOTNOŚĆ GLEBY WILGOTNOŚĆ GLEBY'
   Button "Button_8" at 496,125 size 65x40; TextOff '+ / +2%'
      on Click: function_dd21b452("Wilgotnosc_gleby_auto", 2)
   Button "Button_9" at 497,177 size 65x40; TextOff '- / -2%'
      on Click: function_b9b71300("Wilgotnosc_gleby_auto", 2)
   IOField "I/O field_5" at 508,276 size 62x40; FormatPattern 999
      ProcessValue <- "Wilgotnosc_gleby_auto"
   IOField "I/O field_6" at 508,346 size 62x40; FormatPattern 999
      ProcessValue <- "Czujnik_wilgotności_gleby"
   TextField "Text field_12" at 493,264 size 101x22; Text 'USTAWIONA'
   TextField "Text field_13" at 497,335 size 86x22; Text 'AKTUALNA'
   TextField "Text field_14" at 547,285 size 23x22; Text '%'
   TextField "Text field_15" at 547,356 size 23x22; Text '%'
   Button "Button_10" at 298,125 size 65x40; TextOff '+ / +5%'
      on Click: function_dd21b452("Wilgotnosc_powietrza_auto", 5)
   Button "Button_11" at 298,177 size 65x40; TextOff '- / -5%'
      on Click: function_b9b71300("Wilgotnosc_powietrza_auto", 5)
   IOField "I/O field_4" at 305,277 size 66x40; FormatPattern 999
      ProcessValue <- "Wilgotnosc_powietrza_auto"
   IOField "I/O field_7" at 307,349 size 62x40; FormatPattern 999
      ProcessValue <- "Czujnik_wilgotności_powietrza"
   TextField "Text field_16" at 292,264 size 101x22; Text 'USTAWIONA'
   TextField "Text field_17" at 294,335 size 86x22; Text 'AKTUALNA'
   TextField "Text field_18" at 346,286 size 23x22; Text '%'
   TextField "Text field_19" at 346,357 size 23x22; Text '%'
   Button "Button_14" at 3,1 size 43x43; TextOff 'DOM'; PictureOff "home_1"
      on Click: ActivateScreen("Root screen", 0)
   TextField "Text field_4" at 38,424 size 128x23; Text 'SYSTEM OKIEN'
   Switch "Switch_1" at 198,418 size 185x35; TextOn 'ON'; CaptionText 'Switch'; TextOff 'OFF'
      ProcessValue <- "System_okien_auto"
   GraphicView "Graphic view_1" at 150,60 size 40x40; Picture "Thermometer_icon"
   GraphicView "Graphic view_2" at 330,61 size 40x40; Picture "sensor_4212519"
   TextField "Text field_5" at 93,334 size 86x22; Text 'AKTUALNA'
   TextField "Text field_6" at 90,262 size 101x22; Text 'USTAWIONA'
   GraphicView "Graphic view_3" at 526,61 size 40x40; Picture "soil-sensor_11298794"
   TextField "Text field_1" at 250,4 size 288x34; Text 'TRYB AUTOMATYCZNY'
   Bar "Bar_3" at 620,105 size 70x275; MinimumValue 0; MaximumValue 1500
      ProcessValue <- "Naslonecznienie_auto"
   TextField "Text field_7" at 604,53 size 161x42; Text 'WOLGOTNOŚĆ GLEBY NASŁONECZNIENIE'
   GraphicView "Graphic view_4" at 725,79 size 40x40; Picture "sensor_4212513"
   Button "Button_4" at 696,125 size 65x40; TextOff '+ +50 W m'
      on Click: function_dd21b452("Naslonecznienie_auto", 50)
   Button "Button_5" at 697,177 size 65x40; TextOff '- -50 W m'
      on Click: function_b9b71300("Naslonecznienie_auto", 50)
   IOField "I/O field_3" at 708,276 size 62x40; FormatPattern 999
      ProcessValue <- "Naslonecznienie_auto"
   TextField "Text field_8" at 693,264 size 101x22; Text 'USTAWIONA'
   IOField "I/O field_8" at 711,347 size 62x40; FormatPattern 999
      ProcessValue <- "Czujnik_natezenia_światła"
   TextField "Text field_20" at 697,335 size 86x22; Text 'AKTUALNA'
   TextField "Text field_21" at 747,285 size 23x22; Text '%'
   TextField "Text field_22" at 747,356 size 23x22; Text '%'
   TextField "Text field_23" at 751,143 size 32x18; Text '2'
   TextField "Text field_24" at 748,196 size 32x18; Text '2'

Template "Template_1" 800x480
   Button "Exit" at 671,429 size 71x50; TextOn 'Exit'; TextOff 'Exit'; PictureOn "ExitRuntime_KTP700_Basic_PN_TR"; PictureOff "ExitRuntime_KTP700_Basic_PN_TR"
      on Release: StopRuntime(0)
   Button "Alarms" at 524,429 size 71x50; TextOn 'Alarms'; TextOff 'Alarms'; PictureOn "AlarmDisplay_KTP700_Basic_PN_TR"; PictureOff "AlarmDisplay_KTP700_Basic_PN_TR"
      on Release: function_ef3f5d25("Alarm window_Unacknowledged", -1)
   Button "Start screen" at 169,429 size 71x50; TextOn 'Start screen'; TextOff 'Start screen'; PictureOn "NavigateHome_KTP700_Basic_PN_TR"; PictureOff "NavigateHome_KTP700_Basic_PN_TR"
      on Release: ActivateScreen("Root screen", 0)
      Visibility <- "AlwaysTRUE"
   Button "Language" at 377,429 size 71x50; TextOn 'Language'; TextOff 'Language'; PictureOn "ToggleLanguage_KTP700_Basic_PN_TR"; PictureOff "ToggleLanguage_KTP700_Basic_PN_TR"
      on Release: function_fb9197e8(-1)
*)